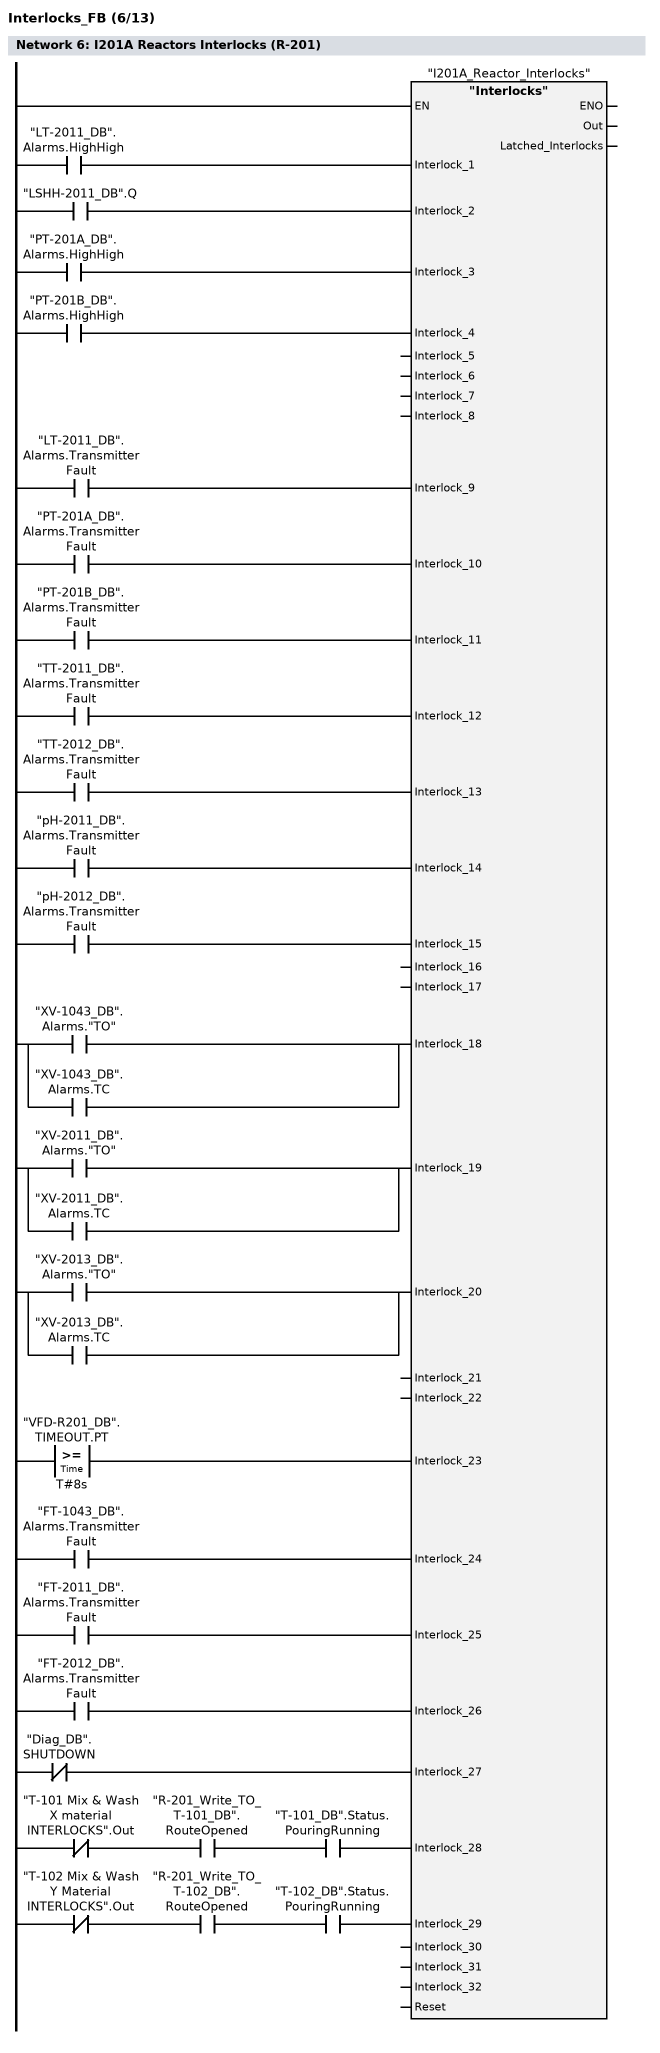
   RUNG wire#powerrail
      "I201A_Reactor_Interlocks"(Interlock_1 := wire#w1, Interlock_2 := wire#w2, Interlock_3 := wire#w3, Interlock_4 := wire#w4, Interlock_9 := wire#w5, Interlock_10 := wire#w6, Interlock_11 := wire#w7, Interlock_12 := wire#w8, Interlock_13 := wire#w9, Interlock_14 := wire#w10, Interlock_15 := wire#w11, Interlock_18 := wire#w12, Interlock_19 := wire#w13, Interlock_20 := wire#w14, Interlock_23 := wire#w15, Interlock_24 := wire#w16, Interlock_25 := wire#w17, Interlock_26 := wire#w18, Interlock_27 := wire#w19, Interlock_28 := wire#w20, Interlock_29 := wire#w21, Interlock_5 :=, Interlock_6 :=, Interlock_7 :=, Interlock_8 :=, Interlock_16 :=, Interlock_17 :=, Interlock_21 :=, Interlock_22 :=, Interlock_30 :=, Interlock_31 :=, Interlock_32 :=, Reset :=, Out =>, Latched_Interlocks =>)
   END_RUNG
   RUNG wire#powerrail
      Contact( "LT-2011_DB".Alarms.HighHigh )
   END_RUNG wire#w1
   RUNG wire#powerrail
      Contact( "LSHH-2011_DB".Q )
   END_RUNG wire#w2
   RUNG wire#powerrail
      Contact( "PT-201A_DB".Alarms.HighHigh )
   END_RUNG wire#w3
   RUNG wire#powerrail
      Contact( "PT-201B_DB".Alarms.HighHigh )
   END_RUNG wire#w4
   RUNG wire#powerrail
      Contact( "LT-2011_DB".Alarms.TransmitterFault )
   END_RUNG wire#w5
   RUNG wire#powerrail
      Contact( "PT-201A_DB".Alarms.TransmitterFault )
   END_RUNG wire#w6
   RUNG wire#powerrail
      Contact( "PT-201B_DB".Alarms.TransmitterFault )
   END_RUNG wire#w7
   RUNG wire#powerrail
      Contact( "TT-2011_DB".Alarms.TransmitterFault )
   END_RUNG wire#w8
   RUNG wire#powerrail
      Contact( "TT-2012_DB".Alarms.TransmitterFault )
   END_RUNG wire#w9
   RUNG wire#powerrail
      Contact( "pH-2011_DB".Alarms.TransmitterFault )
   END_RUNG wire#w10
   RUNG wire#powerrail
      Contact( "pH-2012_DB".Alarms.TransmitterFault )
   END_RUNG wire#w11
   RUNG wire#powerrail
      Contact( "XV-1043_DB".Alarms."TO" )
   END_RUNG wire#w12
   RUNG wire#powerrail
      Contact( "XV-1043_DB".Alarms.TC )
   END_RUNG wire#w12
   RUNG wire#powerrail
      Contact( "XV-2011_DB".Alarms."TO" )
   END_RUNG wire#w13
   RUNG wire#powerrail
      Contact( "XV-2011_DB".Alarms.TC )
   END_RUNG wire#w13
   RUNG wire#powerrail
      Contact( "XV-2013_DB".Alarms."TO" )
   END_RUNG wire#w14
   RUNG wire#powerrail
      Contact( "XV-2013_DB".Alarms.TC )
   END_RUNG wire#w14
   RUNG wire#powerrail
      { S7_Templates := "SrcType := Time" } GE_Contact(in1 := "VFD-R201_DB".TIMEOUT.PT, in2 := T#8s)
   END_RUNG wire#w15
   RUNG wire#powerrail
      Contact( "FT-1043_DB".Alarms.TransmitterFault )
   END_RUNG wire#w16
   RUNG wire#powerrail
      Contact( "FT-2011_DB".Alarms.TransmitterFault )
   END_RUNG wire#w17
   RUNG wire#powerrail
      Contact( "FT-2012_DB".Alarms.TransmitterFault )
   END_RUNG wire#w18
   RUNG wire#powerrail
      I_Contact( "Diag_DB".SHUTDOWN )
   END_RUNG wire#w19
   RUNG wire#powerrail
      I_Contact( "T-101 Mix & Wash X material INTERLOCKS".Out )
      Contact( "R-201_Write_TO_T-101_DB".RouteOpened )
      Contact( "T-101_DB".Status.PouringRunning )
   END_RUNG wire#w20
   RUNG wire#powerrail
      I_Contact( "T-102 Mix & Wash Y Material  INTERLOCKS".Out )
      Contact( "R-201_Write_TO_T-102_DB".RouteOpened )
      Contact( "T-102_DB".Status.PouringRunning )
   END_RUNG wire#w21
   // the same network as SCL:
   "I201A_Reactor_Interlocks"(Interlock_1 := "LT-2011_DB".Alarms.HighHigh,   // "Interlocks"
                           Interlock_2 := "LSHH-2011_DB".Q,
                           Interlock_3 := "PT-201A_DB".Alarms.HighHigh,
                           Interlock_4 := "PT-201B_DB".Alarms.HighHigh,
                           Interlock_9 := "LT-2011_DB".Alarms.TransmitterFault,
                           Interlock_10 := "PT-201A_DB".Alarms.TransmitterFault,
                           Interlock_11 := "PT-201B_DB".Alarms.TransmitterFault,
                           Interlock_12 := "TT-2011_DB".Alarms.TransmitterFault,
                           Interlock_13 := "TT-2012_DB".Alarms.TransmitterFault,
                           Interlock_14 := "pH-2011_DB".Alarms.TransmitterFault,
                           Interlock_15 := "pH-2012_DB".Alarms.TransmitterFault,
                           Interlock_18 := "XV-1043_DB".Alarms."TO" OR "XV-1043_DB".Alarms.TC,
                           Interlock_19 := "XV-2011_DB".Alarms."TO" OR "XV-2011_DB".Alarms.TC,
                           Interlock_20 := "XV-2013_DB".Alarms."TO" OR "XV-2013_DB".Alarms.TC,
                           Interlock_23 := "VFD-R201_DB".TIMEOUT.PT >= T#8s,
                           Interlock_24 := "FT-1043_DB".Alarms.TransmitterFault,
                           Interlock_25 := "FT-2011_DB".Alarms.TransmitterFault,
                           Interlock_26 := "FT-2012_DB".Alarms.TransmitterFault,
                           Interlock_27 := NOT "Diag_DB".SHUTDOWN,
                           Interlock_28 := NOT "T-101 Mix & Wash X material INTERLOCKS".Out AND "R-201_Write_TO_T-101_DB".RouteOpened AND "T-101_DB".Status.PouringRunning,
                           Interlock_29 := NOT "T-102 Mix & Wash Y Material  INTERLOCKS".Out AND "R-201_Write_TO_T-102_DB".RouteOpened AND "T-102_DB".Status.PouringRunning);
END_REGION

REGION Network 7: I201B Reactors Interlocks
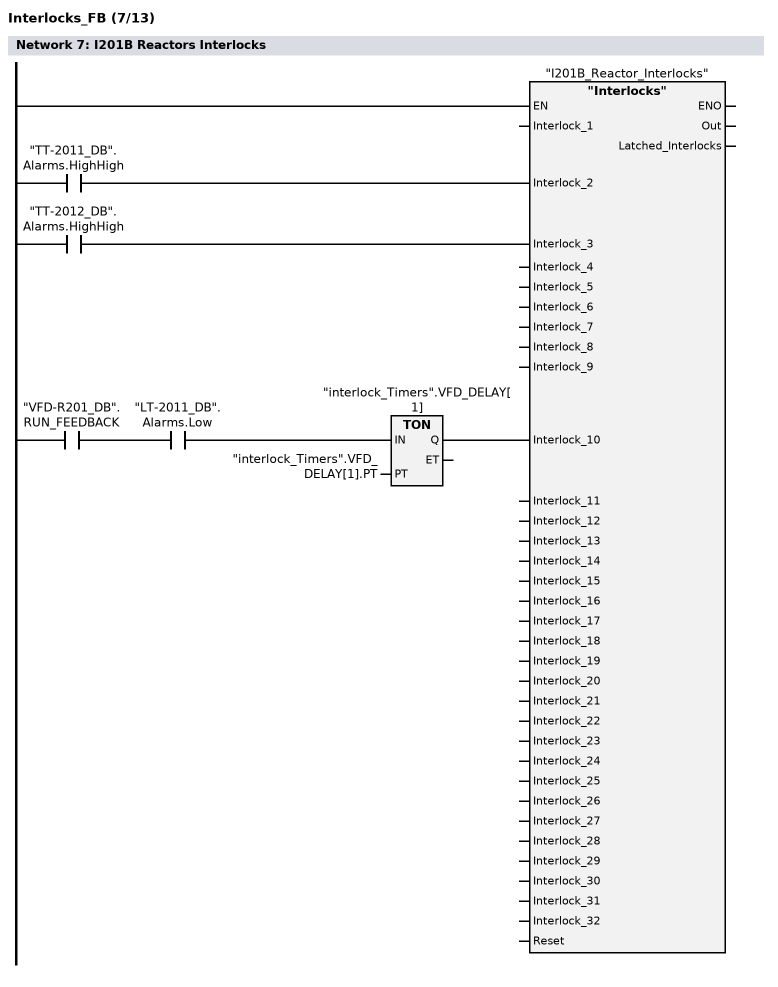
   "interlock_Timers".VFD_DELAY[1].TON(IN := "VFD-R201_DB".RUN_FEEDBACK AND "LT-2011_DB".Alarms.Low,
                           PT := "interlock_Timers".VFD_DELAY[1].PT);
   "I201B_Reactor_Interlocks"(Interlock_2 := "TT-2011_DB".Alarms.HighHigh,   // "Interlocks"
                           Interlock_3 := "TT-2012_DB".Alarms.HighHigh,
                           Interlock_10 := "interlock_Timers".VFD_DELAY[1].Q);
END_REGION

REGION Network 8: I202A Reactors Interlocks
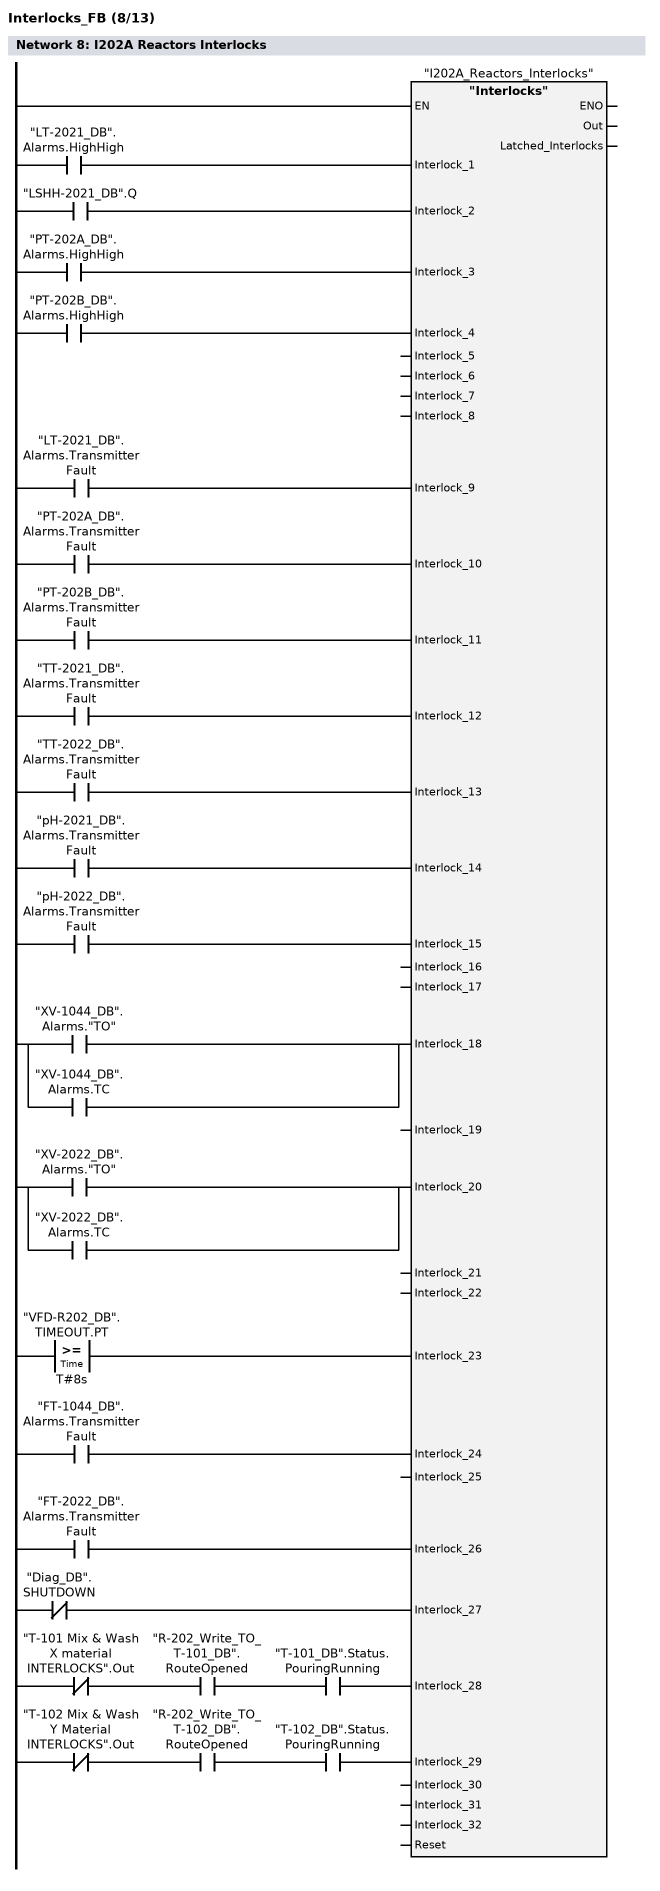
   RUNG wire#powerrail
      "I202A_Reactors_Interlocks"(Interlock_1 := wire#w1, Interlock_2 := wire#w2, Interlock_3 := wire#w3, Interlock_4 := wire#w4, Interlock_9 := wire#w5, Interlock_10 := wire#w6, Interlock_11 := wire#w7, Interlock_12 := wire#w8, Interlock_13 := wire#w9, Interlock_14 := wire#w10, Interlock_15 := wire#w11, Interlock_18 := wire#w12, Interlock_20 := wire#w13, Interlock_23 := wire#w14, Interlock_24 := wire#w15, Interlock_26 := wire#w16, Interlock_27 := wire#w17, Interlock_28 := wire#w18, Interlock_29 := wire#w19, Interlock_5 :=, Interlock_6 :=, Interlock_7 :=, Interlock_8 :=, Interlock_16 :=, Interlock_17 :=, Interlock_19 :=, Interlock_21 :=, Interlock_22 :=, Interlock_25 :=, Interlock_30 :=, Interlock_31 :=, Interlock_32 :=, Reset :=, Out =>, Latched_Interlocks =>)
   END_RUNG
   RUNG wire#powerrail
      Contact( "LT-2021_DB".Alarms.HighHigh )
   END_RUNG wire#w1
   RUNG wire#powerrail
      Contact( "LSHH-2021_DB".Q )
   END_RUNG wire#w2
   RUNG wire#powerrail
      Contact( "PT-202A_DB".Alarms.HighHigh )
   END_RUNG wire#w3
   RUNG wire#powerrail
      Contact( "PT-202B_DB".Alarms.HighHigh )
   END_RUNG wire#w4
   RUNG wire#powerrail
      Contact( "LT-2021_DB".Alarms.TransmitterFault )
   END_RUNG wire#w5
   RUNG wire#powerrail
      Contact( "PT-202A_DB".Alarms.TransmitterFault )
   END_RUNG wire#w6
   RUNG wire#powerrail
      Contact( "PT-202B_DB".Alarms.TransmitterFault )
   END_RUNG wire#w7
   RUNG wire#powerrail
      Contact( "TT-2021_DB".Alarms.TransmitterFault )
   END_RUNG wire#w8
   RUNG wire#powerrail
      Contact( "TT-2022_DB".Alarms.TransmitterFault )
   END_RUNG wire#w9
   RUNG wire#powerrail
      Contact( "pH-2021_DB".Alarms.TransmitterFault )
   END_RUNG wire#w10
   RUNG wire#powerrail
      Contact( "pH-2022_DB".Alarms.TransmitterFault )
   END_RUNG wire#w11
   RUNG wire#powerrail
      Contact( "XV-1044_DB".Alarms."TO" )
   END_RUNG wire#w12
   RUNG wire#powerrail
      Contact( "XV-1044_DB".Alarms.TC )
   END_RUNG wire#w12
   RUNG wire#powerrail
      Contact( "XV-2022_DB".Alarms."TO" )
   END_RUNG wire#w13
   RUNG wire#powerrail
      Contact( "XV-2022_DB".Alarms.TC )
   END_RUNG wire#w13
   RUNG wire#powerrail
      { S7_Templates := "SrcType := Time" } GE_Contact(in1 := "VFD-R202_DB".TIMEOUT.PT, in2 := T#8s)
   END_RUNG wire#w14
   RUNG wire#powerrail
      Contact( "FT-1044_DB".Alarms.TransmitterFault )
   END_RUNG wire#w15
   RUNG wire#powerrail
      Contact( "FT-2022_DB".Alarms.TransmitterFault )
   END_RUNG wire#w16
   RUNG wire#powerrail
      I_Contact( "Diag_DB".SHUTDOWN )
   END_RUNG wire#w17
   RUNG wire#powerrail
      I_Contact( "T-101 Mix & Wash X material INTERLOCKS".Out )
      Contact( "R-202_Write_TO_T-101_DB".RouteOpened )
      Contact( "T-101_DB".Status.PouringRunning )
   END_RUNG wire#w18
   RUNG wire#powerrail
      I_Contact( "T-102 Mix & Wash Y Material  INTERLOCKS".Out )
      Contact( "R-202_Write_TO_T-102_DB".RouteOpened )
      Contact( "T-102_DB".Status.PouringRunning )
   END_RUNG wire#w19
   // the same network as SCL:
   "I202A_Reactors_Interlocks"(Interlock_1 := "LT-2021_DB".Alarms.HighHigh,   // "Interlocks"
                           Interlock_2 := "LSHH-2021_DB".Q,
                           Interlock_3 := "PT-202A_DB".Alarms.HighHigh,
                           Interlock_4 := "PT-202B_DB".Alarms.HighHigh,
                           Interlock_9 := "LT-2021_DB".Alarms.TransmitterFault,
                           Interlock_10 := "PT-202A_DB".Alarms.TransmitterFault,
                           Interlock_11 := "PT-202B_DB".Alarms.TransmitterFault,
                           Interlock_12 := "TT-2021_DB".Alarms.TransmitterFault,
                           Interlock_13 := "TT-2022_DB".Alarms.TransmitterFault,
                           Interlock_14 := "pH-2021_DB".Alarms.TransmitterFault,
                           Interlock_15 := "pH-2022_DB".Alarms.TransmitterFault,
                           Interlock_18 := "XV-1044_DB".Alarms."TO" OR "XV-1044_DB".Alarms.TC,
                           Interlock_20 := "XV-2022_DB".Alarms."TO" OR "XV-2022_DB".Alarms.TC,
                           Interlock_23 := "VFD-R202_DB".TIMEOUT.PT >= T#8s,
                           Interlock_24 := "FT-1044_DB".Alarms.TransmitterFault,
                           Interlock_26 := "FT-2022_DB".Alarms.TransmitterFault,
                           Interlock_27 := NOT "Diag_DB".SHUTDOWN,
                           Interlock_28 := NOT "T-101 Mix & Wash X material INTERLOCKS".Out AND "R-202_Write_TO_T-101_DB".RouteOpened AND "T-101_DB".Status.PouringRunning,
                           Interlock_29 := NOT "T-102 Mix & Wash Y Material  INTERLOCKS".Out AND "R-202_Write_TO_T-102_DB".RouteOpened AND "T-102_DB".Status.PouringRunning);
END_REGION

REGION Network 9: I202B Reactors Interlocks
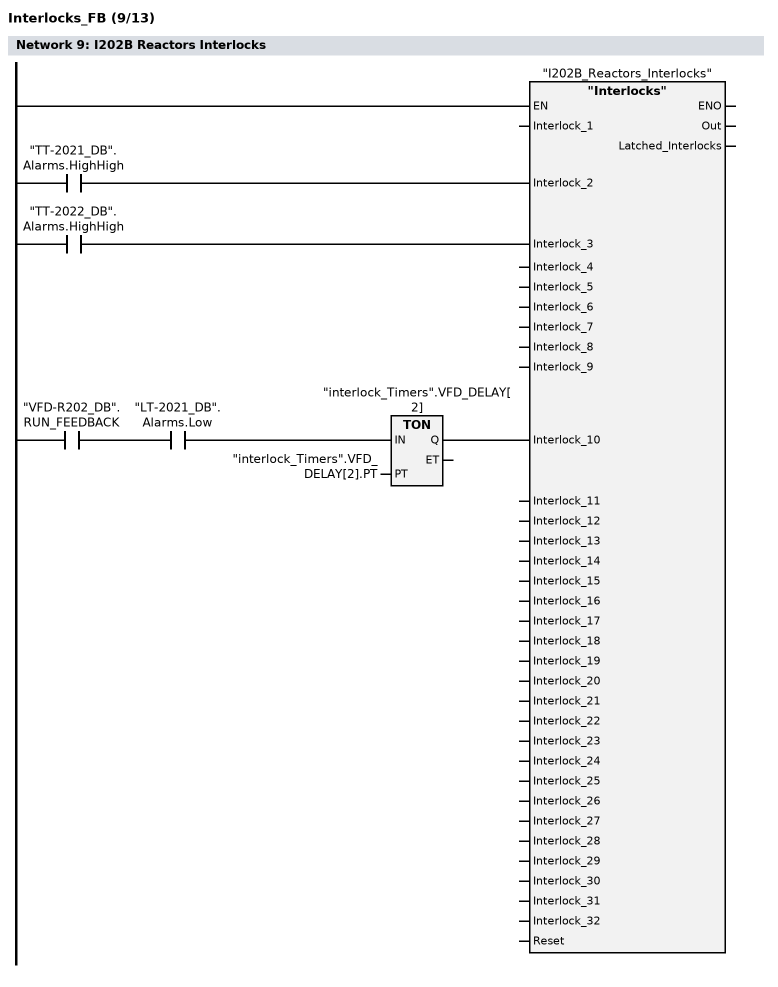
   "interlock_Timers".VFD_DELAY[2].TON(IN := "VFD-R202_DB".RUN_FEEDBACK AND "LT-2021_DB".Alarms.Low,
                           PT := "interlock_Timers".VFD_DELAY[2].PT);
   "I202B_Reactors_Interlocks"(Interlock_2 := "TT-2021_DB".Alarms.HighHigh,   // "Interlocks"
                           Interlock_3 := "TT-2022_DB".Alarms.HighHigh,
                           Interlock_10 := "interlock_Timers".VFD_DELAY[2].Q);
END_REGION

REGION Network 10: I103A Reactor Interlocks
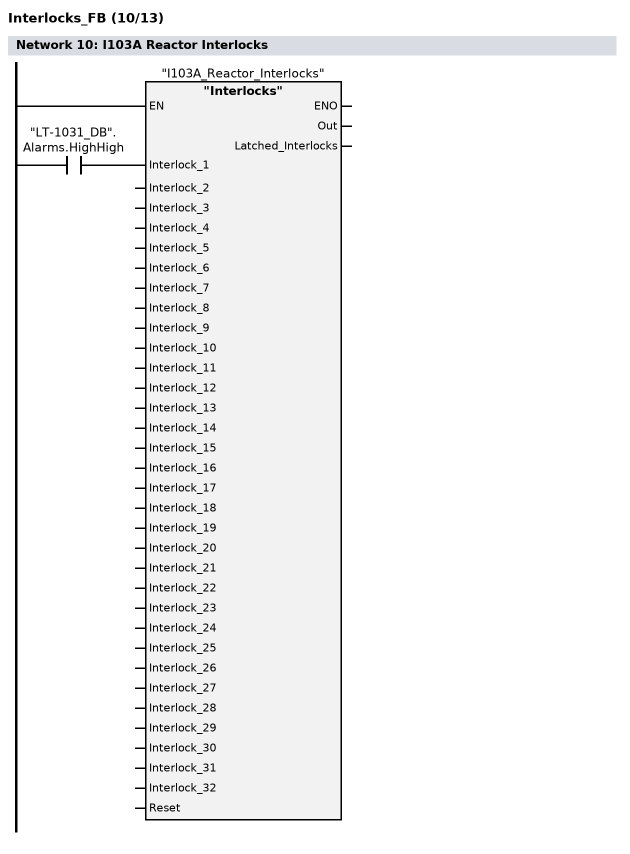
   RUNG wire#powerrail
      "I103A_Reactor_Interlocks"(Interlock_1 := wire#w1, Interlock_2 :=, Interlock_3 :=, Interlock_4 :=, Interlock_5 :=, Interlock_6 :=, Interlock_7 :=, Interlock_8 :=, Interlock_9 :=, Interlock_10 :=, Interlock_11 :=, Interlock_12 :=, Interlock_13 :=, Interlock_14 :=, Interlock_15 :=, Interlock_16 :=, Interlock_17 :=, Interlock_18 :=, Interlock_19 :=, Interlock_20 :=, Interlock_21 :=, Interlock_22 :=, Interlock_23 :=, Interlock_24 :=, Interlock_25 :=, Interlock_26 :=, Interlock_27 :=, Interlock_28 :=, Interlock_29 :=, Interlock_30 :=, Interlock_31 :=, Interlock_32 :=, Reset :=, Out =>, Latched_Interlocks =>)
   END_RUNG
   RUNG wire#powerrail
      Contact( "LT-1031_DB".Alarms.HighHigh )
   END_RUNG wire#w1
   // the same network as SCL:
   "I103A_Reactor_Interlocks"(Interlock_1 := "LT-1031_DB".Alarms.HighHigh);   // "Interlocks"
END_REGION

REGION Network 11: I103B Reactor Interlocks
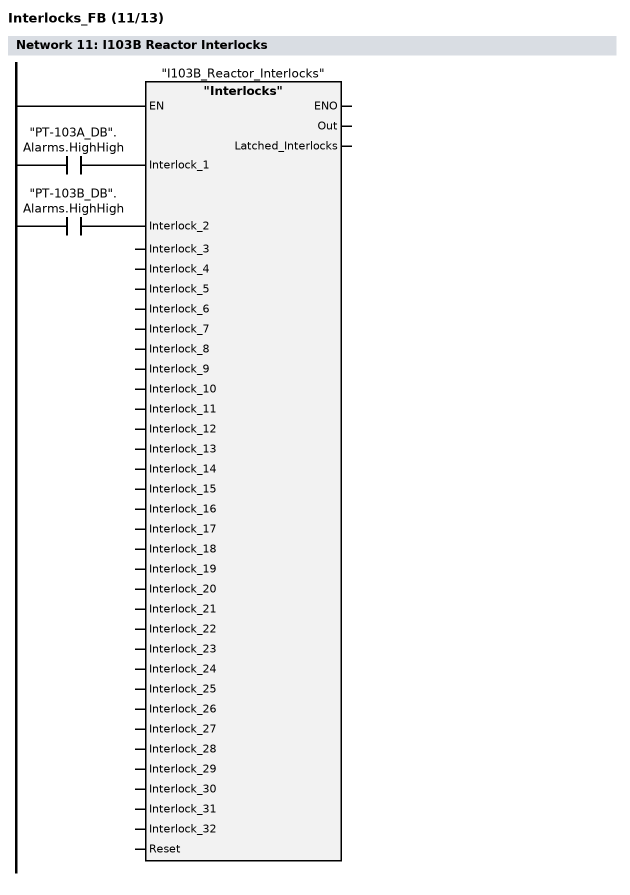
   RUNG wire#powerrail
      "I103B_Reactor_Interlocks"(Interlock_1 := wire#w1, Interlock_2 := wire#w2, Interlock_3 :=, Interlock_4 :=, Interlock_5 :=, Interlock_6 :=, Interlock_7 :=, Interlock_8 :=, Interlock_9 :=, Interlock_10 :=, Interlock_11 :=, Interlock_12 :=, Interlock_13 :=, Interlock_14 :=, Interlock_15 :=, Interlock_16 :=, Interlock_17 :=, Interlock_18 :=, Interlock_19 :=, Interlock_20 :=, Interlock_21 :=, Interlock_22 :=, Interlock_23 :=, Interlock_24 :=, Interlock_25 :=, Interlock_26 :=, Interlock_27 :=, Interlock_28 :=, Interlock_29 :=, Interlock_30 :=, Interlock_31 :=, Interlock_32 :=, Reset :=, Out =>, Latched_Interlocks =>)
   END_RUNG
   RUNG wire#powerrail
      Contact( "PT-103A_DB".Alarms.HighHigh )
   END_RUNG wire#w1
   RUNG wire#powerrail
      Contact( "PT-103B_DB".Alarms.HighHigh )
   END_RUNG wire#w2
   // the same network as SCL:
   "I103B_Reactor_Interlocks"(Interlock_1 := "PT-103A_DB".Alarms.HighHigh,   // "Interlocks"
                           Interlock_2 := "PT-103B_DB".Alarms.HighHigh);
END_REGION

REGION Network 12: I103C Reactor Interlocks
   // Diagnostics for analog output for VFD-1031, VFD-
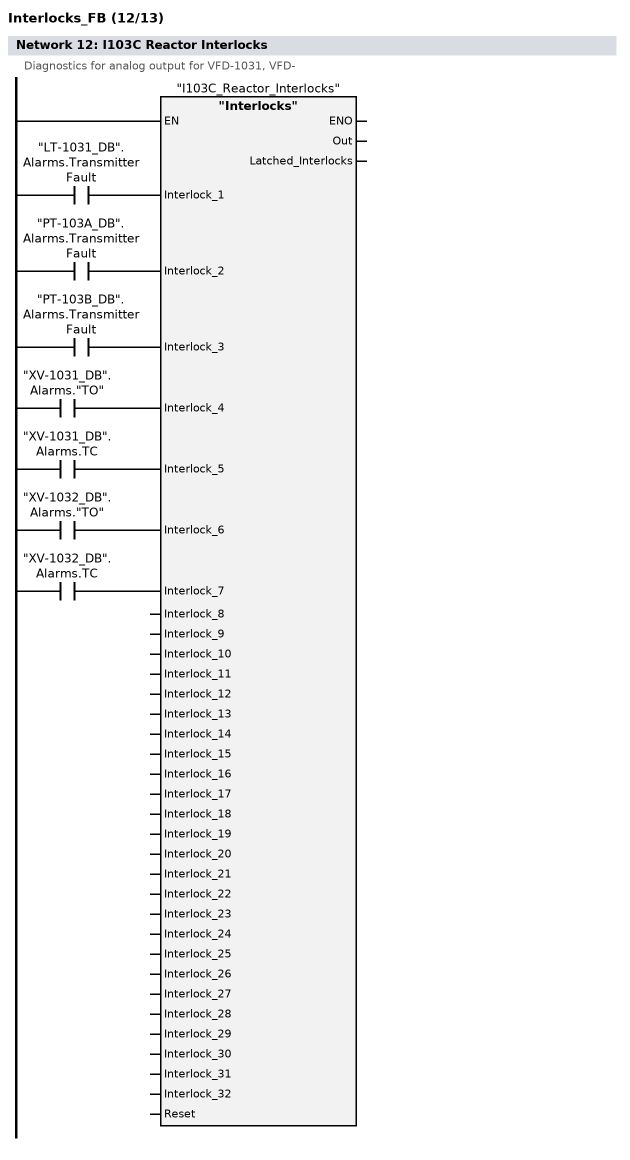
   RUNG wire#powerrail
      "I103C_Reactor_Interlocks"(Interlock_1 := wire#w1, Interlock_2 := wire#w2, Interlock_3 := wire#w3, Interlock_4 := wire#w4, Interlock_5 := wire#w5, Interlock_6 := wire#w6, Interlock_7 := wire#w7, Interlock_8 :=, Interlock_9 :=, Interlock_10 :=, Interlock_11 :=, Interlock_12 :=, Interlock_13 :=, Interlock_14 :=, Interlock_15 :=, Interlock_16 :=, Interlock_17 :=, Interlock_18 :=, Interlock_19 :=, Interlock_20 :=, Interlock_21 :=, Interlock_22 :=, Interlock_23 :=, Interlock_24 :=, Interlock_25 :=, Interlock_26 :=, Interlock_27 :=, Interlock_28 :=, Interlock_29 :=, Interlock_30 :=, Interlock_31 :=, Interlock_32 :=, Reset :=, Out =>, Latched_Interlocks =>)
   END_RUNG
   RUNG wire#powerrail
      Contact( "LT-1031_DB".Alarms.TransmitterFault )
   END_RUNG wire#w1
   RUNG wire#powerrail
      Contact( "PT-103A_DB".Alarms.TransmitterFault )
   END_RUNG wire#w2
   RUNG wire#powerrail
      Contact( "PT-103B_DB".Alarms.TransmitterFault )
   END_RUNG wire#w3
   RUNG wire#powerrail
      Contact( "XV-1031_DB".Alarms."TO" )
   END_RUNG wire#w4
   RUNG wire#powerrail
      Contact( "XV-1031_DB".Alarms.TC )
   END_RUNG wire#w5
   RUNG wire#powerrail
      Contact( "XV-1032_DB".Alarms."TO" )
   END_RUNG wire#w6
   RUNG wire#powerrail
      Contact( "XV-1032_DB".Alarms.TC )
   END_RUNG wire#w7
   // the same network as SCL:
   "I103C_Reactor_Interlocks"(Interlock_1 := "LT-1031_DB".Alarms.TransmitterFault,   // "Interlocks"
                           Interlock_2 := "PT-103A_DB".Alarms.TransmitterFault,
                           Interlock_3 := "PT-103B_DB".Alarms.TransmitterFault,
                           Interlock_4 := "XV-1031_DB".Alarms."TO",
                           Interlock_5 := "XV-1031_DB".Alarms.TC,
                           Interlock_6 := "XV-1032_DB".Alarms."TO",
                           Interlock_7 := "XV-1032_DB".Alarms.TC);
END_REGION

REGION Network 13: I103D Reacotor Interlocks
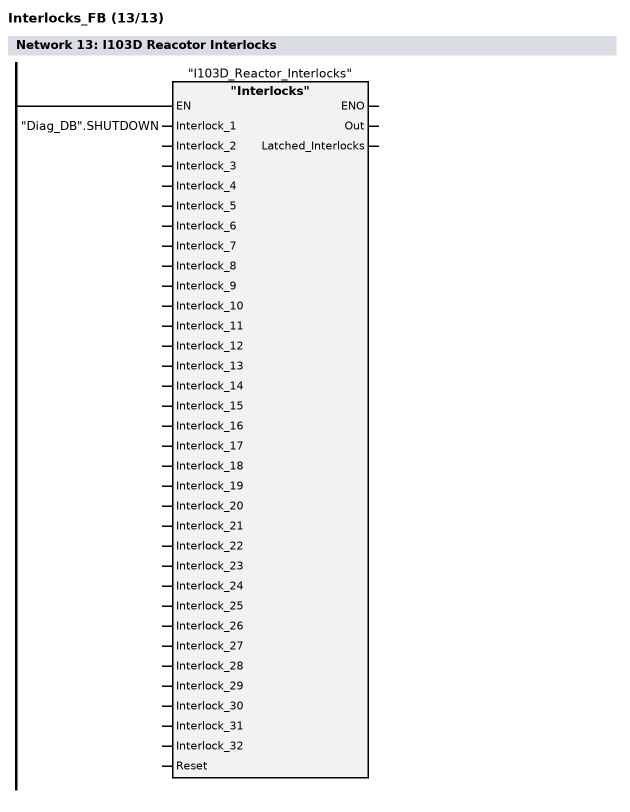
   RUNG wire#powerrail
      "I103D_Reactor_Interlocks"(Interlock_1 := "Diag_DB".SHUTDOWN, Interlock_2 :=, Interlock_3 :=, Interlock_4 :=, Interlock_5 :=, Interlock_6 :=, Interlock_7 :=, Interlock_8 :=, Interlock_9 :=, Interlock_10 :=, Interlock_11 :=, Interlock_12 :=, Interlock_13 :=, Interlock_14 :=, Interlock_15 :=, Interlock_16 :=, Interlock_17 :=, Interlock_18 :=, Interlock_19 :=, Interlock_20 :=, Interlock_21 :=, Interlock_22 :=, Interlock_23 :=, Interlock_24 :=, Interlock_25 :=, Interlock_26 :=, Interlock_27 :=, Interlock_28 :=, Interlock_29 :=, Interlock_30 :=, Interlock_31 :=, Interlock_32 :=, Reset :=, Out =>, Latched_Interlocks =>)
   END_RUNG
   // the same network as SCL:
   "I103D_Reactor_Interlocks"(Interlock_1 := "Diag_DB".SHUTDOWN);   // "Interlocks"
END_REGION
END_FUNCTION

FUNCTION "Interlocks_As_Units" : Void   // FC35, LAD
{ S7_Optimized_Access := 'TRUE' }
VERSION : 0.1
   VAR_TEMP   // added for the SCL form of the ladder/FBD networks
      _w1 : Bool;
   END_VAR
BEGIN

REGION Network 1: R-201 as Unit Interlocks
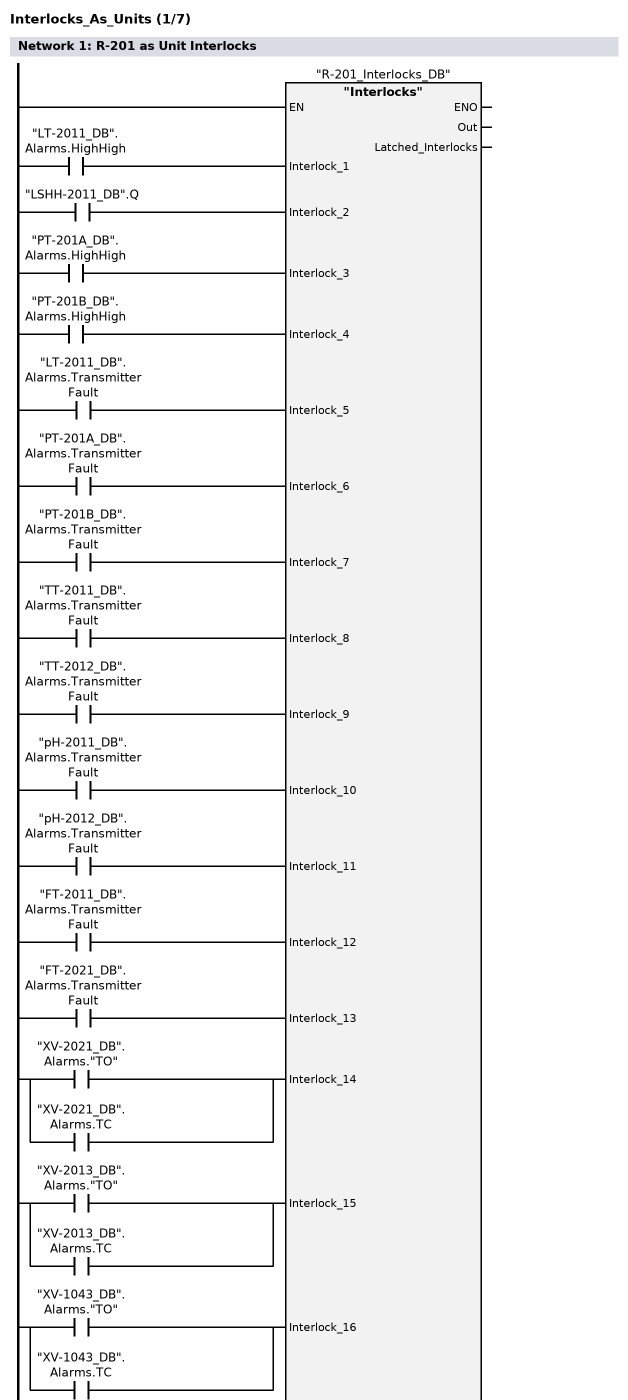
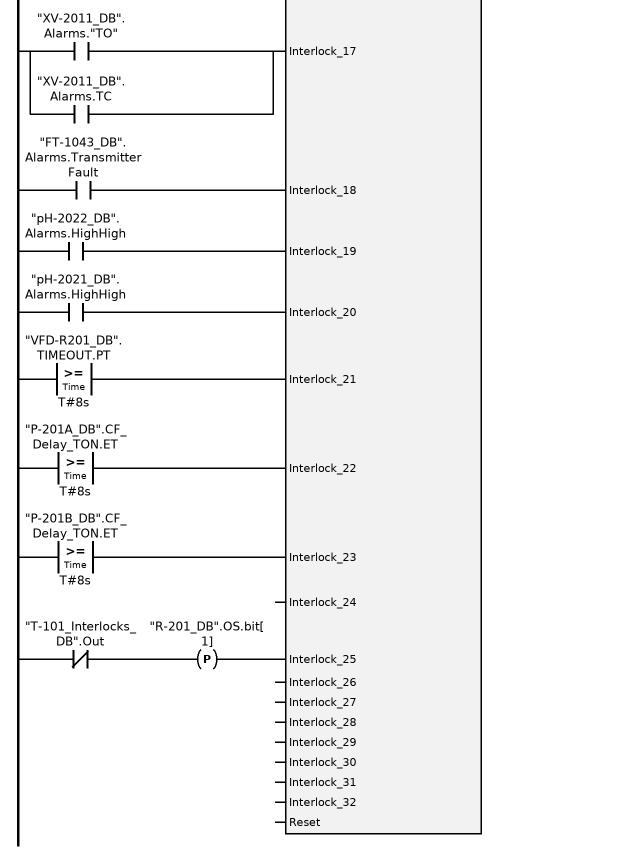
   RUNG wire#powerrail
      "R-201_Interlocks_DB"(Interlock_1 := wire#w1, Interlock_2 := wire#w2, Interlock_3 := wire#w3, Interlock_4 := wire#w4, Interlock_5 := wire#w5, Interlock_6 := wire#w6, Interlock_7 := wire#w7, Interlock_8 := wire#w8, Interlock_9 := wire#w9, Interlock_10 := wire#w10, Interlock_11 := wire#w11, Interlock_12 := wire#w12, Interlock_13 := wire#w13, Interlock_14 := wire#w14, Interlock_15 := wire#w15, Interlock_16 := wire#w16, Interlock_17 := wire#w17, Interlock_18 := wire#w18, Interlock_19 := wire#w19, Interlock_20 := wire#w20, Interlock_21 := wire#w21, Interlock_22 := wire#w22, Interlock_23 := wire#w23, Interlock_25 := wire#w24, Interlock_24 :=, Interlock_26 :=, Interlock_27 :=, Interlock_28 :=, Interlock_29 :=, Interlock_30 :=, Interlock_31 :=, Interlock_32 :=, Reset :=, Out =>, Latched_Interlocks =>)
   END_RUNG
   RUNG wire#powerrail
      Contact( "LT-2011_DB".Alarms.HighHigh )
   END_RUNG wire#w1
   RUNG wire#powerrail
      Contact( "LSHH-2011_DB".Q )
   END_RUNG wire#w2
   RUNG wire#powerrail
      Contact( "PT-201A_DB".Alarms.HighHigh )
   END_RUNG wire#w3
   RUNG wire#powerrail
      Contact( "PT-201B_DB".Alarms.HighHigh )
   END_RUNG wire#w4
   RUNG wire#powerrail
      Contact( "LT-2011_DB".Alarms.TransmitterFault )
   END_RUNG wire#w5
   RUNG wire#powerrail
      Contact( "PT-201A_DB".Alarms.TransmitterFault )
   END_RUNG wire#w6
   RUNG wire#powerrail
      Contact( "PT-201B_DB".Alarms.TransmitterFault )
   END_RUNG wire#w7
   RUNG wire#powerrail
      Contact( "TT-2011_DB".Alarms.TransmitterFault )
   END_RUNG wire#w8
   RUNG wire#powerrail
      Contact( "TT-2012_DB".Alarms.TransmitterFault )
   END_RUNG wire#w9
   RUNG wire#powerrail
      Contact( "pH-2011_DB".Alarms.TransmitterFault )
   END_RUNG wire#w10
   RUNG wire#powerrail
      Contact( "pH-2012_DB".Alarms.TransmitterFault )
   END_RUNG wire#w11
   RUNG wire#powerrail
      Contact( "FT-2011_DB".Alarms.TransmitterFault )
   END_RUNG wire#w12
   RUNG wire#powerrail
      Contact( "FT-2021_DB".Alarms.TransmitterFault )
   END_RUNG wire#w13
   RUNG wire#powerrail
      Contact( "XV-2021_DB".Alarms."TO" )
   END_RUNG wire#w14
   RUNG wire#powerrail
      Contact( "XV-2021_DB".Alarms.TC )
   END_RUNG wire#w14
   RUNG wire#powerrail
      Contact( "XV-2013_DB".Alarms."TO" )
   END_RUNG wire#w15
   RUNG wire#powerrail
      Contact( "XV-2013_DB".Alarms.TC )
   END_RUNG wire#w15
   RUNG wire#powerrail
      Contact( "XV-1043_DB".Alarms."TO" )
   END_RUNG wire#w16
   RUNG wire#powerrail
      Contact( "XV-1043_DB".Alarms.TC )
   END_RUNG wire#w16
   RUNG wire#powerrail
      Contact( "XV-2011_DB".Alarms."TO" )
   END_RUNG wire#w17
   RUNG wire#powerrail
      Contact( "XV-2011_DB".Alarms.TC )
   END_RUNG wire#w17
   RUNG wire#powerrail
      Contact( "FT-1043_DB".Alarms.TransmitterFault )
   END_RUNG wire#w18
   RUNG wire#powerrail
      Contact( "pH-2022_DB".Alarms.HighHigh )
   END_RUNG wire#w19